
           //------------------------------------------------------------------------------------------
           // Convert relative to absoulte coordinates
           //------------------------------------------------------------------------------------------
           // check for additional circMode = 3 to be activated (LKinLang)
           // Changes CmdType to absolute and converts cirmode 3 to 1
           // --> CmdType = 3 (always absolute as result)
           // --> CircleParameters = calculated arc & updated auxPoint
           IF #pathDataElementPreBuf.cmdParameters.circleParameters.circMode = "LKINCTRL_CIRCMODE_GCODE"
             AND #statSubfunctionStatus = #STATUS_NO_ERROR
           THEN
             #tempRetValWord := "LKinCtrl_ConvCircMode3To1"(coordinates := #pathDataElementPreBuf.cmdCoordinates.absolutePosition,
                                                            lastPos := #statLastPos,
                                                            errorMessage => #statDebugMessage,
                                                            cmdType := #pathDataElementPreBuf.cmdType,
                                                            circleParameters := #pathDataElementPreBuf.cmdParameters.circleParameters);
           END_IF;

           IF #statSubfunctionStatus = #STATUS_NO_ERROR THEN
             // Calculate resulting absoulte position; also convert relative to absolute positions
             #tempRetValWord := "LKinCtrl_CalcResultingPos"(cmdType := #pathDataElementPreBuf.cmdType,
                                                            cartesianPos := #pathDataElementPreBuf.cmdCoordinates.absolutePosition,
                                                            circleParameters := #pathDataElementPreBuf.cmdParameters.circleParameters,
                                                            errorMessage => #statDebugMessage,
                                                            lastAuxPoint := #statAuxPoint, // Absoulte auxPoint
                                                            lastPos := #statLastPos); // Absolute endPoint

             // After this FC call the lastPos equals the endPoint and absolute position
             #statEndPoint := #statAbsolutePosition := #statLastPos;

             // Check if ResultingPos calculation returned an error
             IF #tempRetValWord <> #STATUS_NO_ERROR THEN
               // set error information
               #diagnostics.faultSetNumber := #pathDataElementPreBuf.cmdID;
               #diagnostics.faultPathDataName := #pathDataElementPreBuf.pathDataName;
               #statSubfunctionStatus := #tempRetValWord;
               // set state machine
               #statStateMachine := #ERROR_STATE;
             END_IF;
           END_IF;

         ELSE
           // Command is not a motion command --> WaitTime or FlagOnly
           // ==> Nothing to calculate 
           ;
         END_IF;

         //------------------------------------------------------------------------------------------
         // Command Selection
         //------------------------------------------------------------------------------------------
         // interpretation command to be a linear or circular motion
         IF #statSubfunctionStatus = #STATUS_NO_ERROR THEN
           IF #pathDataElementPreBuf.cmdType = "LKINCTRL_MC_MOVELINEARABS" OR
             #pathDataElementPreBuf.cmdType = "LKINCTRL_MC_MOVELINEARREL" THEN
             #statStateMachine := #EXEC_LIN;
           ELSIF #pathDataElementPreBuf.cmdType = "LKINCTRL_MC_MOVECIRCULARABS" OR
             #pathDataElementPreBuf.cmdType = "LKINCTRL_MC_MOVECIRCULARREL" THEN
             #statStateMachine := #EXEC_CIRC;
           ELSIF #pathDataElementPreBuf.cmdType = "LKINCTRL_MC_MOVEDIRECTABS" OR
             #pathDataElementPreBuf.cmdType = "LKINCTRL_MC_MOVEDIRECTREL" THEN
             #statStateMachine := #EXEC_MOVE_DIRECT;
           ELSIF #pathDataElementPreBuf.cmdType = "LKINCTRL_CMD_WAIT_TIME" THEN
             #statStateMachine := #EXEC_WAIT_TIME;
           ELSIF #pathDataElementPreBuf.cmdType = "LKINCTRL_CMD_FLAG_ONLY" THEN
             #statStateMachine := #EXEC_FLAG_ONLY;
           ELSIF #pathDataElementPreBuf.cmdType = "LKINCTRL_MC_TRACKCONVEYORBELT" THEN
             #statStateMachine := #EXEC_TRACK_CONV;
           END_IF;
         END_IF;
       END_IF;

     END_REGION CMD_CALC 


     // execute MC_MOVELINEARABSOLUTE motion commands  
     REGION EXEC_LIN
       IF #statStateMachine = #EXEC_LIN
         // AND #statDebugState = TRUE
       THEN
         // reset  variable for single step debugging of states
         #statDebugState := FALSE;

         IF #statError = FALSE THEN

           // set execute trigger for linear command
           #statExecLinCmds[#statFBCounterLin] := TRUE;

           // Store motion command data for further calcualtions
           // last position for relative commands
           //#statLastPos := #statAbsolutePosition;

           // command details from PathData and assignment to MC_FBs for activeCmdNo
           #statStoreExecuteBuffer.bufferElement[#statStoreExecuteBuffer.writeBufferElement].pathDataName := #pathDataElementPreBuf.pathDataName;
           #statStoreExecuteBuffer.bufferElement[#statStoreExecuteBuffer.writeBufferElement].pathDataIdentifier := #pathDataElementPreBuf.pathDataIdentifier;
           #statStoreExecuteBuffer.bufferElement[#statStoreExecuteBuffer.writeBufferElement].setNumber := #pathDataElementPreBuf.cmdID;
           #statStoreExecuteBuffer.bufferElement[#statStoreExecuteBuffer.writeBufferElement].MotionFBNo := #statFBCounterLin;
           #statStoreExecuteBuffer.lastBufferElement := #statStoreExecuteBuffer.writeBufferElement;

           // increase writeBufferElement pointer for statStoreBuffer for assignment of activeCmdNo
           IF #statStoreExecuteBuffer.writeBufferElement < #LKINCTRL_EXECUTEBUFFER_LENGTH THEN
             #statStoreExecuteBuffer.writeBufferElement := #statStoreExecuteBuffer.writeBufferElement + 1;
           ELSE
             #statStoreExecuteBuffer.writeBufferElement := 1;
           END_IF;

           REGION CMD_LOGGER
             // // DATA LOGGER handling
             // write command data to data logger
             // single data entries of PathDataElement instead of complete structure ==> to deep nesting level
             #statDebugExecCmdLogger.loggerElement[#statDebugExecCmdLogger.writeCmdLoggerElement].executedCmd.cmdType := #pathDataElementPreBuf.cmdType;
             #statDebugExecCmdLogger.loggerElement[#statDebugExecCmdLogger.writeCmdLoggerElement].executedCmd.pathDataName := #pathDataElementPreBuf.pathDataName;
             #statDebugExecCmdLogger.loggerElement[#statDebugExecCmdLogger.writeCmdLoggerElement].executedCmd.pathDataIdentifier := #pathDataElementPreBuf.pathDataIdentifier;
             #statDebugExecCmdLogger.loggerElement[#statDebugExecCmdLogger.writeCmdLoggerElement].executedCmd.cmdID := #pathDataElementPreBuf.cmdID;
             #statDebugExecCmdLogger.loggerElement[#statDebugExecCmdLogger.writeCmdLoggerElement].executedCmd.cmdName := #pathDataElementPreBuf.cmdName;
             // coordinates logging
             #statDebugExecCmdLogger.loggerElement[#statDebugExecCmdLogger.writeCmdLoggerElement].executedCmd.coordinateX := #pathDataElementPreBuf.cmdCoordinates.absolutePosition[1];
             #statDebugExecCmdLogger.loggerElement[#statDebugExecCmdLogger.writeCmdLoggerElement].executedCmd.coordinateY := #pathDataElementPreBuf.cmdCoordinates.absolutePosition[2];
             #statDebugExecCmdLogger.loggerElement[#statDebugExecCmdLogger.writeCmdLoggerElement].executedCmd.coordinateZ := #pathDataElementPreBuf.cmdCoordinates.absolutePosition[3];
             #statDebugExecCmdLogger.loggerElement[#statDebugExecCmdLogger.writeCmdLoggerElement].executedCmd.coordinateA := #pathDataElementPreBuf.cmdCoordinates.absolutePosition[4];
             #statDebugExecCmdLogger.loggerElement[#statDebugExecCmdLogger.writeCmdLoggerElement].executedCmd.coordSystem := #pathDataElementPreBuf.cmdCoordinates.coordSystem;
             // cmdParameter logging
             #statDebugExecCmdLogger.loggerElement[#statDebugExecCmdLogger.writeCmdLoggerElement].executedCmd.bufferMode := #pathDataElementPreBuf.cmdParameters.bufferMode;
             #statDebugExecCmdLogger.loggerElement[#statDebugExecCmdLogger.writeCmdLoggerElement].executedCmd.transitionParameter := #pathDataElementPreBuf.cmdParameters.transitionParameters[1];
             #statDebugExecCmdLogger.loggerElement[#statDebugExecCmdLogger.writeCmdLoggerElement].executedCmd.dynVelocity := #pathDataElementPreBuf.cmdParameters.pathDynamics.velocity;
             #statDebugExecCmdLogger.loggerElement[#statDebugExecCmdLogger.writeCmdLoggerElement].executedCmd.dynAcceleration := #pathDataElementPreBuf.cmdParameters.pathDynamics.acceleration;
             #statDebugExecCmdLogger.loggerElement[#statDebugExecCmdLogger.writeCmdLoggerElement].executedCmd.dynDeceleration := #pathDataElementPreBuf.cmdParameters.pathDynamics.deceleration;
             #statDebugExecCmdLogger.loggerElement[#statDebugExecCmdLogger.writeCmdLoggerElement].executedCmd.dynJerk := #pathDataElementPreBuf.cmdParameters.pathDynamics.jerk;
             #statDebugExecCmdLogger.loggerElement[#statDebugExecCmdLogger.writeCmdLoggerElement].executedCmd.dynamicAdpation := #pathDataElementPreBuf.cmdParameters.dynamicAdaption;
             // logger element data
             #statDebugExecCmdLogger.loggerElement[#statDebugExecCmdLogger.writeCmdLoggerElement].executeBufferElement := #statStoreExecuteBuffer.lastBufferElement;
             #statDebugExecCmdLogger.loggerElement[#statDebugExecCmdLogger.writeCmdLoggerElement].assignedMotionFB := #statFBCounterLin;
             #tempRetVal := RD_SYS_T(#statDebugExecCmdLogger.loggerElement[#statDebugExecCmdLogger.writeCmdLoggerElement].timeStamp);

             // increment writeCmdLogger pointer
             IF #statDebugExecCmdLogger.writeCmdLoggerElement < #CONST_LENGTH_DATALOGGER THEN
               #statDebugExecCmdLogger.writeCmdLoggerElement := #statDebugExecCmdLogger.writeCmdLoggerElement + 1;
             ELSE
               #statDebugExecCmdLogger.writeCmdLoggerElement := 1;
             END_IF;
           END_REGION CMD_LOGGER

           // set FBCounter variables
           IF #statFBCounterLin < #LKINCTRL_MAX_NUMBER_OF_CMDS_LIN THEN
             #statFBCounterLin := #statFBCounterLin + 1;
           ELSE
             #statFBCounterLin := 1;
           END_IF;

           // set status for outputs
           #statCmdExecuted := TRUE;
           #statStatus := #STATUS_CMD_EXECUTED;

         ELSE
           #statStateMachine := #ERROR_STATE;
         END_IF;
       END_IF;
     END_REGION EXEC_LIN


     // execute MC_MOVECIRCULRABSOLUTE motion commands
     REGION EXEC_CIRC
       IF #statStateMachine = #EXEC_CIRC
         // AND #statDebugState = TRUE
       THEN
         // reset variable for single step debugging of states
         #statDebugState := FALSE;

         IF #statError = FALSE THEN

           // set execute trigger for circular command
           #statExecCircCmds[#statFBCounterCirc] := TRUE;

           // command details from PathData and assignment to MC_FBs for activeCmdNo
           #statStoreExecuteBuffer.bufferElement[#statStoreExecuteBuffer.writeBufferElement].pathDataName := #pathDataElementPreBuf.pathDataName;
           #statStoreExecuteBuffer.bufferElement[#statStoreExecuteBuffer.writeBufferElement].pathDataIdentifier := #pathDataElementPreBuf.pathDataIdentifier;
           #statStoreExecuteBuffer.bufferElement[#statStoreExecuteBuffer.writeBufferElement].setNumber := #pathDataElementPreBuf.cmdID;
           #statStoreExecuteBuffer.bufferElement[#statStoreExecuteBuffer.writeBufferElement].MotionFBNo := #LKINCTRL_EXECUTEBUFFER_LENGTH + #statFBCounterCirc;
           #statStoreExecuteBuffer.lastBufferElement := #statStoreExecuteBuffer.writeBufferElement;

           // increase writeBufferElement pointer for statStoreBuffer for assignment of activeCmdNo
           IF #statStoreExecuteBuffer.writeBufferElement < #LKINCTRL_EXECUTEBUFFER_LENGTH THEN
             #statStoreExecuteBuffer.writeBufferElement := #statStoreExecuteBuffer.writeBufferElement + 1;
           ELSE
             #statStoreExecuteBuffer.writeBufferElement := 1;
           END_IF;

           REGION CMD_LOGGER
             // // DATA LOGGER handling
             // write command data to data logger
             // single data entries of PathDataElement instead of complete structure ==> to deep nesting level
             #statDebugExecCmdLogger.loggerElement[#statDebugExecCmdLogger.writeCmdLoggerElement].executedCmd.cmdType := #pathDataElementPreBuf.cmdType;
             #statDebugExecCmdLogger.loggerElement[#statDebugExecCmdLogger.writeCmdLoggerElement].executedCmd.pathDataName := #pathDataElementPreBuf.pathDataName;
             #statDebugExecCmdLogger.loggerElement[#statDebugExecCmdLogger.writeCmdLoggerElement].executedCmd.pathDataIdentifier := #pathDataElementPreBuf.pathDataIdentifier;
             #statDebugExecCmdLogger.loggerElement[#statDebugExecCmdLogger.writeCmdLoggerElement].executedCmd.cmdID := #pathDataElementPreBuf.cmdID;
             #statDebugExecCmdLogger.loggerElement[#statDebugExecCmdLogger.writeCmdLoggerElement].executedCmd.cmdName := #pathDataElementPreBuf.cmdName;
             // coordinates logging (use auxPoint in X,Y,Z variables)
             #statDebugExecCmdLogger.loggerElement[#statDebugExecCmdLogger.writeCmdLoggerElement].executedCmd.coordinateX := #statEndPoint[1];
             #statDebugExecCmdLogger.loggerElement[#statDebugExecCmdLogger.writeCmdLoggerElement].executedCmd.coordinateY := #statEndPoint[2];
             #statDebugExecCmdLogger.loggerElement[#statDebugExecCmdLogger.writeCmdLoggerElement].executedCmd.coordinateZ := #statEndPoint[3];
             #statDebugExecCmdLogger.loggerElement[#statDebugExecCmdLogger.writeCmdLoggerElement].executedCmd.coordinateA := #statEndPoint[4];
             #statDebugExecCmdLogger.loggerElement[#statDebugExecCmdLogger.writeCmdLoggerElement].executedCmd.coordSystem := #pathDataElementPreBuf.cmdCoordinates.coordSystem;
             // cmdParameter logging
             #statDebugExecCmdLogger.loggerElement[#statDebugExecCmdLogger.writeCmdLoggerElement].executedCmd.bufferMode := #pathDataElementPreBuf.cmdParameters.bufferMode;
             #statDebugExecCmdLogger.loggerElement[#statDebugExecCmdLogger.writeCmdLoggerElement].executedCmd.transitionParameter := #pathDataElementPreBuf.cmdParameters.transitionParameters[1];
             #statDebugExecCmdLogger.loggerElement[#statDebugExecCmdLogger.writeCmdLoggerElement].executedCmd.dynVelocity := #pathDataElementPreBuf.cmdParameters.pathDynamics.velocity;
             #statDebugExecCmdLogger.loggerElement[#statDebugExecCmdLogger.writeCmdLoggerElement].executedCmd.dynAcceleration := #pathDataElementPreBuf.cmdParameters.pathDynamics.acceleration;
             #statDebugExecCmdLogger.loggerElement[#statDebugExecCmdLogger.writeCmdLoggerElement].executedCmd.dynDeceleration := #pathDataElementPreBuf.cmdParameters.pathDynamics.deceleration;
             #statDebugExecCmdLogger.loggerElement[#statDebugExecCmdLogger.writeCmdLoggerElement].executedCmd.dynJerk := #pathDataElementPreBuf.cmdParameters.pathDynamics.jerk;
             #statDebugExecCmdLogger.loggerElement[#statDebugExecCmdLogger.writeCmdLoggerElement].executedCmd.dynamicAdpation := #pathDataElementPreBuf.cmdParameters.dynamicAdaption;
             // circle parameter logging
             #statDebugExecCmdLogger.loggerElement[#statDebugExecCmdLogger.writeCmdLoggerElement].executedCmd.circMode := #pathDataElementPreBuf.cmdParameters.circleParameters.circMode;
             #statDebugExecCmdLogger.loggerElement[#statDebugExecCmdLogger.writeCmdLoggerElement].executedCmd.auxPoint_1 := #pathDataElementPreBuf.cmdParameters.circleParameters.auxPoint[1];
             #statDebugExecCmdLogger.loggerElement[#statDebugExecCmdLogger.writeCmdLoggerElement].executedCmd.auxPoint_2 := #pathDataElementPreBuf.cmdParameters.circleParameters.auxPoint[2];
             #statDebugExecCmdLogger.loggerElement[#statDebugExecCmdLogger.writeCmdLoggerElement].executedCmd.auxPoint_3 := #pathDataElementPreBuf.cmdParameters.circleParameters.auxPoint[3];
             #statDebugExecCmdLogger.loggerElement[#statDebugExecCmdLogger.writeCmdLoggerElement].executedCmd.pathChoice := #pathDataElementPreBuf.cmdParameters.circleParameters.pathChoice;
             #statDebugExecCmdLogger.loggerElement[#statDebugExecCmdLogger.writeCmdLoggerElement].executedCmd.circlePlane := #pathDataElementPreBuf.cmdParameters.circleParameters.circlePlane;
             #statDebugExecCmdLogger.loggerElement[#statDebugExecCmdLogger.writeCmdLoggerElement].executedCmd.radius := #pathDataElementPreBuf.cmdParameters.circleParameters.radius;
             #statDebugExecCmdLogger.loggerElement[#statDebugExecCmdLogger.writeCmdLoggerElement].executedCmd.arc := #pathDataElementPreBuf.cmdParameters.circleParameters.arc;

             // logger element data
             #statDebugExecCmdLogger.loggerElement[#statDebugExecCmdLogger.writeCmdLoggerElement].executeBufferElement := #statStoreExecuteBuffer.lastBufferElement;
             #statDebugExecCmdLogger.loggerElement[#statDebugExecCmdLogger.writeCmdLoggerElement].assignedMotionFB := 10 + #statFBCounterCirc;
             #tempRetVal := RD_SYS_T(#statDebugExecCmdLogger.loggerElement[#statDebugExecCmdLogger.writeCmdLoggerElement].timeStamp);

             // increment writeCmdLogger pointer
             IF #statDebugExecCmdLogger.writeCmdLoggerElement < #CONST_LENGTH_DATALOGGER THEN
               #statDebugExecCmdLogger.writeCmdLoggerElement := #statDebugExecCmdLogger.writeCmdLoggerElement + 1;
             ELSE
               #statDebugExecCmdLogger.writeCmdLoggerElement := 1;
             END_IF;
           END_REGION CMD_LOGGER

           // set FBCounter variables
           IF #statFBCounterCirc < #LKINCTRL_MAX_NUMBER_OF_CMDS_CIRC THEN
             #statFBCounterCirc := #statFBCounterCirc + 1;
           ELSE
             #statFBCounterCirc := 1;
           END_IF;

           // set status for outputs
           #statCmdExecuted := TRUE;
           #statStatus := #STATUS_CMD_EXECUTED;

         ELSE
           #statStateMachine := #ERROR_STATE;
         END_IF;
       END_IF;
     END_REGION EXEC_CIRC


     // execute MC_MOVEDIRECTABSOLUTE motion commands  
     REGION EXEC_MOVE_DIRECT
       IF #statStateMachine = #EXEC_MOVE_DIRECT
         // AND #statDebugState = TRUE
       THEN
         // reset  variable for single step debugging of states
         #statDebugState := FALSE;

         IF #statError = FALSE THEN

           // set execute trigger for move direct command
           #statExecMoveDirectCmds[#statFBCounterMoveDir] := TRUE;

           // Store motion command data for further calcualtions
           // last position for relative commands
           //#statLastPos := #statAbsolutePosition;

           // command details from PathData and assignment to MC_FBs for activeCmdNo
           #statStoreExecuteBuffer.bufferElement[#statStoreExecuteBuffer.writeBufferElement].pathDataName := #pathDataElementPreBuf.pathDataName;
           #statStoreExecuteBuffer.bufferElement[#statStoreExecuteBuffer.writeBufferElement].pathDataIdentifier := #pathDataElementPreBuf.pathDataIdentifier;
           #statStoreExecuteBuffer.bufferElement[#statStoreExecuteBuffer.writeBufferElement].setNumber := #pathDataElementPreBuf.cmdID;
           #statStoreExecuteBuffer.bufferElement[#statStoreExecuteBuffer.writeBufferElement].MotionFBNo := #LKINCTRL_EXECUTEBUFFER_LENGTH + #LKINCTRL_EXECUTEBUFFER_LENGTH + #statFBCounterMoveDir;
           #statStoreExecuteBuffer.lastBufferElement := #statStoreExecuteBuffer.writeBufferElement;

           // increase writeBufferElement pointer for statStoreBuffer for assignment of activeCmdNo
           IF #statStoreExecuteBuffer.writeBufferElement < #LKINCTRL_EXECUTEBUFFER_LENGTH THEN
             #statStoreExecuteBuffer.writeBufferElement := #statStoreExecuteBuffer.writeBufferElement + 1;
           ELSE
             #statStoreExecuteBuffer.writeBufferElement := 1;
           END_IF;

           REGION CMD_LOGGER
             // // DATA LOGGER handling
             // write command data to data logger
             // single data entries of PathDataElement instead of complete structure ==> to deep nesting level
             #statDebugExecCmdLogger.loggerElement[#statDebugExecCmdLogger.writeCmdLoggerElement].executedCmd.cmdType := #pathDataElementPreBuf.cmdType;
             #statDebugExecCmdLogger.loggerElement[#statDebugExecCmdLogger.writeCmdLoggerElement].executedCmd.pathDataName := #pathDataElementPreBuf.pathDataName;
             #statDebugExecCmdLogger.loggerElement[#statDebugExecCmdLogger.writeCmdLoggerElement].executedCmd.pathDataIdentifier := #pathDataElementPreBuf.pathDataIdentifier;
             #statDebugExecCmdLogger.loggerElement[#statDebugExecCmdLogger.writeCmdLoggerElement].executedCmd.cmdID := #pathDataElementPreBuf.cmdID;
             #statDebugExecCmdLogger.loggerElement[#statDebugExecCmdLogger.writeCmdLoggerElement].executedCmd.cmdName := #pathDataElementPreBuf.cmdName;
             // coordinates logging
             #statDebugExecCmdLogger.loggerElement[#statDebugExecCmdLogger.writeCmdLoggerElement].executedCmd.coordinateX := #pathDataElementPreBuf.cmdCoordinates.absolutePosition[1];
             #statDebugExecCmdLogger.loggerElement[#statDebugExecCmdLogger.writeCmdLoggerElement].executedCmd.coordinateY := #pathDataElementPreBuf.cmdCoordinates.absolutePosition[2];
             #statDebugExecCmdLogger.loggerElement[#statDebugExecCmdLogger.writeCmdLoggerElement].executedCmd.coordinateZ := #pathDataElementPreBuf.cmdCoordinates.absolutePosition[3];
             #statDebugExecCmdLogger.loggerElement[#statDebugExecCmdLogger.writeCmdLoggerElement].executedCmd.coordinateA := #pathDataElementPreBuf.cmdCoordinates.absolutePosition[4];
             #statDebugExecCmdLogger.loggerElement[#statDebugExecCmdLogger.writeCmdLoggerElement].executedCmd.coordSystem := #pathDataElementPreBuf.cmdCoordinates.coordSystem;
             // cmdParameter logging
             #statDebugExecCmdLogger.loggerElement[#statDebugExecCmdLogger.writeCmdLoggerElement].executedCmd.bufferMode := #pathDataElementPreBuf.cmdParameters.bufferMode;
             #statDebugExecCmdLogger.loggerElement[#statDebugExecCmdLogger.writeCmdLoggerElement].executedCmd.transitionParameter := #pathDataElementPreBuf.cmdParameters.transitionParameters[1];
             #statDebugExecCmdLogger.loggerElement[#statDebugExecCmdLogger.writeCmdLoggerElement].executedCmd.dynVelocity := #pathDataElementPreBuf.cmdParameters.pathDynamics.velocity;
             #statDebugExecCmdLogger.loggerElement[#statDebugExecCmdLogger.writeCmdLoggerElement].executedCmd.dynAcceleration := #pathDataElementPreBuf.cmdParameters.pathDynamics.acceleration;
             #statDebugExecCmdLogger.loggerElement[#statDebugExecCmdLogger.writeCmdLoggerElement].executedCmd.dynDeceleration := #pathDataElementPreBuf.cmdParameters.pathDynamics.deceleration;
             #statDebugExecCmdLogger.loggerElement[#statDebugExecCmdLogger.writeCmdLoggerElement].executedCmd.dynJerk := #pathDataElementPreBuf.cmdParameters.pathDynamics.jerk;
             #statDebugExecCmdLogger.loggerElement[#statDebugExecCmdLogger.writeCmdLoggerElement].executedCmd.dynamicAdpation := #pathDataElementPreBuf.cmdParameters.dynamicAdaption;

             #statDebugExecCmdLogger.loggerElement[#statDebugExecCmdLogger.writeCmdLoggerElement].executedCmd.linkConstellation := #pathDataElementPreBuf.cmdParameters.moveDirectParameters.linkConstellation;
             #statDebugExecCmdLogger.loggerElement[#statDebugExecCmdLogger.writeCmdLoggerElement].executedCmd.positionMode := #pathDataElementPreBuf.cmdParameters.moveDirectParameters.positionMode;

             // logger element data
             #statDebugExecCmdLogger.loggerElement[#statDebugExecCmdLogger.writeCmdLoggerElement].executeBufferElement := #statStoreExecuteBuffer.lastBufferElement;
             #statDebugExecCmdLogger.loggerElement[#statDebugExecCmdLogger.writeCmdLoggerElement].assignedMotionFB := #statFBCounterMoveDir;
             #tempRetVal := RD_SYS_T(#statDebugExecCmdLogger.loggerElement[#statDebugExecCmdLogger.writeCmdLoggerElement].timeStamp);

             // increment writeCmdLogger pointer
             IF #statDebugExecCmdLogger.writeCmdLoggerElement < #CONST_LENGTH_DATALOGGER THEN
               #statDebugExecCmdLogger.writeCmdLoggerElement := #statDebugExecCmdLogger.writeCmdLoggerElement + 1;
             ELSE
               #statDebugExecCmdLogger.writeCmdLoggerElement := 1;
             END_IF;
           END_REGION CMD_LOGGER

           // set FBCounter variables
           IF #statFBCounterMoveDir < #LKINCTRL_MAX_NUMBER_OF_CMDS_MOVEDIRECT THEN
             #statFBCounterMoveDir := #statFBCounterMoveDir + 1;
           ELSE
             #statFBCounterMoveDir := 1;
           END_IF;

           // set status for outputs
           #statCmdExecuted := TRUE;
           #statStatus := #STATUS_CMD_EXECUTED;

         ELSE
           #statStateMachine := #ERROR_STATE;
         END_IF;
       END_IF;
     END_REGION EXEC_MOVE_DIRECT


     // execute MC_TRACKCONVEYORBELT motion commands  
     REGION EXEC_TRACK_CONVEYOR
       IF #statStateMachine = #EXEC_TRACK_CONV
         // AND #statDebugState = TRUE
       THEN
         // reset  variable for single step debugging of states
         #statDebugState := FALSE;

         IF #statError = FALSE THEN

           // set execute trigger for move direct command
           #statExecTrackConv[#statFBCounterTrackConv] := TRUE;

           // Copy conveyor configuration to instance
           #statConveyorBeltAxis[#statFBCounterTrackConv] := #conveyorConfiguration[#pathDataElementPreBuf.cmdParameters.conveyorParameters.conveyorParaNo].conveyorBeltAxis;
           #instMC_TrackConveyor[#statFBCounterTrackConv].ConveyorBeltOrigin := #conveyorConfiguration[#pathDataElementPreBuf.cmdParameters.conveyorParameters.conveyorParaNo].conveyorBeltOrigin;
           #instMC_TrackConveyor[#statFBCounterTrackConv].InitialObjectPosition := #conveyorConfiguration[#pathDataElementPreBuf.cmdParameters.conveyorParameters.conveyorParaNo].initialObjectPosition;
           #instMC_TrackConveyor[#statFBCounterTrackConv].CoordSystem := #pathDataElementPreBuf.cmdCoordinates.coordSystem;

           // Set OCS in tracking
           #statOCSInTracking[#instMC_TrackConveyor[#statFBCounterTrackConv].CoordSystem] := TRUE;

           // command details from PathData and assignment to MC_FBs for activeCmdNo
           #statStoreExecuteBuffer.bufferElement[#statStoreExecuteBuffer.writeBufferElement].pathDataName := #pathDataElementPreBuf.pathDataName;
           #statStoreExecuteBuffer.bufferElement[#statStoreExecuteBuffer.writeBufferElement].pathDataIdentifier := #pathDataElementPreBuf.pathDataIdentifier;
           #statStoreExecuteBuffer.bufferElement[#statStoreExecuteBuffer.writeBufferElement].setNumber := #pathDataElementPreBuf.cmdID;
           #statStoreExecuteBuffer.bufferElement[#statStoreExecuteBuffer.writeBufferElement].MotionFBNo := "LKINCTRL_CMD_WAIT_TIME" + #statFBCounterTrackConv;
           #statStoreExecuteBuffer.lastBufferElement := #statStoreExecuteBuffer.writeBufferElement;

           // increase writeBufferElement pointer for statStoreBuffer for assignment of activeCmdNo
           IF #statStoreExecuteBuffer.writeBufferElement < #LKINCTRL_EXECUTEBUFFER_LENGTH THEN
             #statStoreExecuteBuffer.writeBufferElement := #statStoreExecuteBuffer.writeBufferElement + 1;
           ELSE
             #statStoreExecuteBuffer.writeBufferElement := 1;
           END_IF;

           REGION CMD_LOGGER
             // // DATA LOGGER handling
             // write command data to data logger
             // single data entries of PathDataElement instead of complete structure ==> to deep nesting level
             #statDebugExecCmdLogger.loggerElement[#statDebugExecCmdLogger.writeCmdLoggerElement].executedCmd.cmdType := #pathDataElementPreBuf.cmdType;
             #statDebugExecCmdLogger.loggerElement[#statDebugExecCmdLogger.writeCmdLoggerElement].executedCmd.pathDataName := #pathDataElementPreBuf.pathDataName;
             #statDebugExecCmdLogger.loggerElement[#statDebugExecCmdLogger.writeCmdLoggerElement].executedCmd.pathDataIdentifier := #pathDataElementPreBuf.pathDataIdentifier;
             #statDebugExecCmdLogger.loggerElement[#statDebugExecCmdLogger.writeCmdLoggerElement].executedCmd.cmdID := #pathDataElementPreBuf.cmdID;
             #statDebugExecCmdLogger.loggerElement[#statDebugExecCmdLogger.writeCmdLoggerElement].executedCmd.cmdName := #pathDataElementPreBuf.cmdName;
             // coordinates logging
             #statDebugExecCmdLogger.loggerElement[#statDebugExecCmdLogger.writeCmdLoggerElement].executedCmd.coordinateX := #pathDataElementPreBuf.cmdCoordinates.absolutePosition[1];
             #statDebugExecCmdLogger.loggerElement[#statDebugExecCmdLogger.writeCmdLoggerElement].executedCmd.coordinateY := #pathDataElementPreBuf.cmdCoordinates.absolutePosition[2];
             #statDebugExecCmdLogger.loggerElement[#statDebugExecCmdLogger.writeCmdLoggerElement].executedCmd.coordinateZ := #pathDataElementPreBuf.cmdCoordinates.absolutePosition[3];
             #statDebugExecCmdLogger.loggerElement[#statDebugExecCmdLogger.writeCmdLoggerElement].executedCmd.coordinateA := #pathDataElementPreBuf.cmdCoordinates.absolutePosition[4];
             #statDebugExecCmdLogger.loggerElement[#statDebugExecCmdLogger.writeCmdLoggerElement].executedCmd.coordSystem := #pathDataElementPreBuf.cmdCoordinates.coordSystem;
             // cmdParameter logging
             #statDebugExecCmdLogger.loggerElement[#statDebugExecCmdLogger.writeCmdLoggerElement].executedCmd.bufferMode := #pathDataElementPreBuf.cmdParameters.bufferMode;
             #statDebugExecCmdLogger.loggerElement[#statDebugExecCmdLogger.writeCmdLoggerElement].executedCmd.transitionParameter := #pathDataElementPreBuf.cmdParameters.transitionParameters[1];
             #statDebugExecCmdLogger.loggerElement[#statDebugExecCmdLogger.writeCmdLoggerElement].executedCmd.dynVelocity := #pathDataElementPreBuf.cmdParameters.pathDynamics.velocity;
             #statDebugExecCmdLogger.loggerElement[#statDebugExecCmdLogger.writeCmdLoggerElement].executedCmd.dynAcceleration := #pathDataElementPreBuf.cmdParameters.pathDynamics.acceleration;
             #statDebugExecCmdLogger.loggerElement[#statDebugExecCmdLogger.writeCmdLoggerElement].executedCmd.dynDeceleration := #pathDataElementPreBuf.cmdParameters.pathDynamics.deceleration;
             #statDebugExecCmdLogger.loggerElement[#statDebugExecCmdLogger.writeCmdLoggerElement].executedCmd.dynJerk := #pathDataElementPreBuf.cmdParameters.pathDynamics.jerk;
             #statDebugExecCmdLogger.loggerElement[#statDebugExecCmdLogger.writeCmdLoggerElement].executedCmd.dynamicAdpation := #pathDataElementPreBuf.cmdParameters.dynamicAdaption;

             #statDebugExecCmdLogger.loggerElement[#statDebugExecCmdLogger.writeCmdLoggerElement].executedCmd.linkConstellation := #pathDataElementPreBuf.cmdParameters.moveDirectParameters.linkConstellation;
             #statDebugExecCmdLogger.loggerElement[#statDebugExecCmdLogger.writeCmdLoggerElement].executedCmd.positionMode := #pathDataElementPreBuf.cmdParameters.moveDirectParameters.positionMode;

             // logger element data
             #statDebugExecCmdLogger.loggerElement[#statDebugExecCmdLogger.writeCmdLoggerElement].executeBufferElement := #statStoreExecuteBuffer.lastBufferElement;
             #statDebugExecCmdLogger.loggerElement[#statDebugExecCmdLogger.writeCmdLoggerElement].assignedMotionFB := #statFBCounterTrackConv;
             #tempRetVal := RD_SYS_T(#statDebugExecCmdLogger.loggerElement[#statDebugExecCmdLogger.writeCmdLoggerElement].timeStamp);

             // increment writeCmdLogger pointer
             IF #statDebugExecCmdLogger.writeCmdLoggerElement < #CONST_LENGTH_DATALOGGER THEN
               #statDebugExecCmdLogger.writeCmdLoggerElement := #statDebugExecCmdLogger.writeCmdLoggerElement + 1;
             ELSE
               #statDebugExecCmdLogger.writeCmdLoggerElement := 1;
             END_IF;
           END_REGION CMD_LOGGER

           // set FBCounter variables
           IF #statFBCounterTrackConv < #LKINCTRL_MAX_NUMBER_OF_CMDS_TRACKCONV THEN
             #statFBCounterTrackConv := #statFBCounterTrackConv + 1;
           ELSE
             #statFBCounterTrackConv := 1;
           END_IF;

           // set status for outputs
           #statCmdExecuted := TRUE;
           #statStatus := #STATUS_CMD_EXECUTED;

         ELSE
           #statStateMachine := #ERROR_STATE;
         END_IF;
       END_IF;
     END_REGION EXEC_TRACK_CONVEYOR



     // execute WAIT TIME 
     REGION EXEC_WAIT_TIME
       IF #statStateMachine = #EXEC_WAIT_TIME
         // AND #statDebugState = TRUE
       THEN
         // reset  variable for single step debugging of states
         #statDebugState := FALSE;

         // check for error to be pending
         IF #statError = FALSE THEN

           // Added check for active mc command; FR: 27.05.2019
           // check for active MC linear instance
           FOR #tempCtr := 1 TO #LKINCTRL_MAX_NUMBER_OF_CMDS_LIN DO
             IF #instMC_MoveLinAbs[#tempCtr].Busy THEN
               // set temp to interlock reset
               #tempMCActive := TRUE;
               EXIT;
             ELSE
               #tempMCActive := FALSE;
             END_IF;
           END_FOR;

           // check for no circular instance to be busy in case of no linear cmd busy
           IF #tempMCActive = FALSE THEN
             FOR #tempCtr := 1 TO #LKINCTRL_MAX_NUMBER_OF_CMDS_CIRC DO
               IF #instMC_MoveCircAbs[#tempCtr].Busy THEN
                 // set temp to interlock reset
                 #tempMCActive := TRUE;
                 EXIT;
               ELSE
                 #tempMCActive := FALSE;
               END_IF;
             END_FOR;
           END_IF;

           // check for no PTP instance to be busy in case of no linear cmd busy
           IF #tempMCActive = FALSE THEN
             FOR #tempCtr := 1 TO #LKINCTRL_MAX_NUMBER_OF_CMDS_MOVEDIRECT DO
               IF #instMC_MoveDirectAbs[#tempCtr].Busy THEN
                 // set temp to interlock reset
                 #tempMCActive := TRUE;
                 EXIT;
               ELSE
                 #tempMCActive := FALSE;
               END_IF;
             END_FOR;
           END_IF;

           // check for previously executed commands to be finished
           IF #to_Kinematics.StatusMotionQueue.NumberOfCommands = 0
             AND #statActive = FALSE
             AND #tempMCActive = FALSE
           THEN
             // read wait time - duration [ms]
             #statWaitTime := INT_TO_TIME(LREAL_TO_INT(#pathDataElementPreBuf.cmdParameters.pathDynamics.velocity));

             // set execute trigger to run timer
             #statExecWaitTime := TRUE;

             // command details from PathData and assignment to MC_FBs for activeCmdNo
             #statStoreExecuteBuffer.bufferElement[#statStoreExecuteBuffer.writeBufferElement].pathDataName := #pathDataElementPreBuf.pathDataName;
             #statStoreExecuteBuffer.bufferElement[#statStoreExecuteBuffer.writeBufferElement].pathDataIdentifier := #pathDataElementPreBuf.pathDataIdentifier;
             #statStoreExecuteBuffer.bufferElement[#statStoreExecuteBuffer.writeBufferElement].setNumber := #pathDataElementPreBuf.cmdID;
             #statStoreExecuteBuffer.bufferElement[#statStoreExecuteBuffer.writeBufferElement].MotionFBNo := "LKINCTRL_CMD_WAIT_TIME";
             #statStoreExecuteBuffer.lastBufferElement := #statStoreExecuteBuffer.writeBufferElement;

             // increase writeBufferElement pointer for statStoreBuffer for assignment of activeCmdNo
             IF #statStoreExecuteBuffer.writeBufferElement < #LKINCTRL_EXECUTEBUFFER_LENGTH THEN
               #statStoreExecuteBuffer.writeBufferElement := #statStoreExecuteBuffer.writeBufferElement + 1;
             ELSE
               #statStoreExecuteBuffer.writeBufferElement := 1;
             END_IF;

             REGION CMD_LOGGER
               // // DATA LOGGER handling
               // write command data to data logger
               // single data entries of PathDataElement instead of complete structure ==> to deep nesting level
               #statDebugExecCmdLogger.loggerElement[#statDebugExecCmdLogger.writeCmdLoggerElement].executedCmd.cmdType := #pathDataElementPreBuf.cmdType;
               #statDebugExecCmdLogger.loggerElement[#statDebugExecCmdLogger.writeCmdLoggerElement].executedCmd.pathDataName := #pathDataElementPreBuf.pathDataName;
               #statDebugExecCmdLogger.loggerElement[#statDebugExecCmdLogger.writeCmdLoggerElement].executedCmd.pathDataIdentifier := #pathDataElementPreBuf.pathDataIdentifier;
               #statDebugExecCmdLogger.loggerElement[#statDebugExecCmdLogger.writeCmdLoggerElement].executedCmd.cmdID := #pathDataElementPreBuf.cmdID;
               #statDebugExecCmdLogger.loggerElement[#statDebugExecCmdLogger.writeCmdLoggerElement].executedCmd.cmdName := #pathDataElementPreBuf.cmdName;
               // parameter logging
               #statDebugExecCmdLogger.loggerElement[#statDebugExecCmdLogger.writeCmdLoggerElement].executedCmd.dynVelocity := #pathDataElementPreBuf.cmdParameters.pathDynamics.velocity;
               // logger element data
               #statDebugExecCmdLogger.loggerElement[#statDebugExecCmdLogger.writeCmdLoggerElement].executeBufferElement := #statStoreExecuteBuffer.lastBufferElement;
               #statDebugExecCmdLogger.loggerElement[#statDebugExecCmdLogger.writeCmdLoggerElement].assignedMotionFB := "LKINCTRL_CMD_WAIT_TIME";
               #tempRetVal := RD_SYS_T(#statDebugExecCmdLogger.loggerElement[#statDebugExecCmdLogger.writeCmdLoggerElement].timeStamp);

               // increment writeCmdLogger pointer
               IF #statDebugExecCmdLogger.writeCmdLoggerElement < #CONST_LENGTH_DATALOGGER THEN
                 #statDebugExecCmdLogger.writeCmdLoggerElement := #statDebugExecCmdLogger.writeCmdLoggerElement + 1;
               ELSE
                 #statDebugExecCmdLogger.writeCmdLoggerElement := 1;
               END_IF;
             END_REGION CMD_LOGGER

             // set cmdExecuted
             #statCmdExecuted := TRUE;
             // set state to signalize WAIT_TIME running
             #statStatus := #STATUS_WAIT_TIME_ACTIVE;
             // go to state to wait for WAIT_TIME to finish
             #statStateMachine := #WAITING_TIME;
           END_IF;

         ELSE
           #statStateMachine := #ERROR_STATE;
         END_IF;
       END_IF;
     END_REGION EXEC_WAIT_TIME


     // execute FLAG_ONLY commands  
     REGION EXEC_FLAG_ONLY
       IF #statStateMachine = #EXEC_FLAG_ONLY
         // AND #statDebugState = TRUE
       THEN
         // reset  variable for single step debugging of states
         #statDebugState := FALSE;

         IF #statError = FALSE THEN

           // checked for PathData to start with flagOnly command in the triggering section (must not be 1st command)
           // set flagOnlyCmd bit manually, as no previous MC command will be 'done' before

           IF #statStartCmdIsFlagOnly THEN
             // set execute trigger here only when PathData starts with flagOnly command
             #statExecuteFlagOnlyCmd := TRUE;
             // reset bit to recognize FlagOnly command
             #statStartCmdIsFlagOnly := FALSE;
           END_IF;

           // command details from PathData and assignment to MC_FBs for activeCmdNo
           #statStoreExecuteBuffer.bufferElement[#statStoreExecuteBuffer.writeBufferElement].pathDataName := #pathDataElementPreBuf.pathDataName;
           #statStoreExecuteBuffer.bufferElement[#statStoreExecuteBuffer.writeBufferElement].pathDataIdentifier := #pathDataElementPreBuf.pathDataIdentifier;
           #statStoreExecuteBuffer.bufferElement[#statStoreExecuteBuffer.writeBufferElement].setNumber := #pathDataElementPreBuf.cmdID;
           #statStoreExecuteBuffer.bufferElement[#statStoreExecuteBuffer.writeBufferElement].MotionFBNo := "LKINCTRL_CMD_FLAG_ONLY";
           #statStoreExecuteBuffer.lastBufferElement := #statStoreExecuteBuffer.writeBufferElement;

           // increase writeBufferElement pointer for statStoreBuffer for assignment of activeCmdNo
           IF #statStoreExecuteBuffer.writeBufferElement < #LKINCTRL_EXECUTEBUFFER_LENGTH THEN
             #statStoreExecuteBuffer.writeBufferElement := #statStoreExecuteBuffer.writeBufferElement + 1;
           ELSE
             #statStoreExecuteBuffer.writeBufferElement := 1;
           END_IF;

           REGION CMD_LOGGER
             // // DATA LOGGER handling
             // write command data to data logger
             // single data entries of PathDataElement instead of complete structure ==> to deep nesting level
             #statDebugExecCmdLogger.loggerElement[#statDebugExecCmdLogger.writeCmdLoggerElement].executedCmd.cmdType := #pathDataElementPreBuf.cmdType;
             #statDebugExecCmdLogger.loggerElement[#statDebugExecCmdLogger.writeCmdLoggerElement].executedCmd.pathDataName := #pathDataElementPreBuf.pathDataName;
             #statDebugExecCmdLogger.loggerElement[#statDebugExecCmdLogger.writeCmdLoggerElement].executedCmd.pathDataIdentifier := #pathDataElementPreBuf.pathDataIdentifier;
             #statDebugExecCmdLogger.loggerElement[#statDebugExecCmdLogger.writeCmdLoggerElement].executedCmd.cmdID := #pathDataElementPreBuf.cmdID;
             #statDebugExecCmdLogger.loggerElement[#statDebugExecCmdLogger.writeCmdLoggerElement].executedCmd.cmdName := #pathDataElementPreBuf.cmdName;

             // logger element data
             #statDebugExecCmdLogger.loggerElement[#statDebugExecCmdLogger.writeCmdLoggerElement].executeBufferElement := #statStoreExecuteBuffer.lastBufferElement;
             #statDebugExecCmdLogger.loggerElement[#statDebugExecCmdLogger.writeCmdLoggerElement].assignedMotionFB := "LKINCTRL_CMD_FLAG_ONLY";
             #tempRetVal := RD_SYS_T(#statDebugExecCmdLogger.loggerElement[#statDebugExecCmdLogger.writeCmdLoggerElement].timeStamp);

             // increment writeCmdLogger pointer
             IF #statDebugExecCmdLogger.writeCmdLoggerElement < #CONST_LENGTH_DATALOGGER THEN
               #statDebugExecCmdLogger.writeCmdLoggerElement := #statDebugExecCmdLogger.writeCmdLoggerElement + 1;
             ELSE
               #statDebugExecCmdLogger.writeCmdLoggerElement := 1;
             END_IF;
           END_REGION CMD_LOGGER

           // set status for outputs
           #statCmdExecuted := TRUE;
           #statStatus := #STATUS_CMD_EXECUTED;

         ELSE
           #statStateMachine := #ERROR_STATE;
         END_IF;
       END_IF;
     END_REGION EXEC_FLAG_ONLY


     // wait for WAIT_TIME to finish
     REGION WAITING_TIME
       IF #statStateMachine = #WAITING_TIME
         // AND #statDebugState = TRUE
       THEN
         // reset  variable for single step debugging of states
         #statDebugState := FALSE;

         // Set waitTimeActive output
         #statWaitTimeActive := TRUE;

         IF #instIEC_Timer_waitTime.Q THEN
           // reset timer by calling with false
           #statExecWaitTime := FALSE;

           // set status for outputs only after time is done
           #statCmdExecuted := TRUE;

           // Reset output
           #statWaitTimeActive := FALSE;

           #statStatus := #STATUS_WAIT_TIME_FINISHED;
         END_IF;

       END_IF;
     END_REGION WAITING_TIME


     // state reached when GroupInterrupt is interrupted ==> do nothing when interrupted
     REGION CONTINUEING 
       IF #statStateMachine = #CONTINUEING
         // AND #statDebugState = TRUE
       THEN
         // reset  variable for single step debugging of states
         #statDebugState := FALSE;

         // check for MC_GroupContinue to be performed successfully  (TO Kinematics not interrupted anymore)
         IF #to_Kinematics.StatusWord.%X17 = FALSE THEN
           #statStateMachine := #CONTINUED;
         ELSE // Added FR 2019/04/12
           // execute MC_GroupContinue only when kinematics is interrupted
           #statExecGroupContinue := TRUE;
         END_IF;

       END_IF;
     END_REGION CONTINUEING


     // state reached when GroupContinue is done ==> do nothing when path motion continues
     REGION CONTINUED
       IF #statStateMachine = #CONTINUED
         // AND #statDebugState = TRUE
       THEN
         // reset  variable for single step debugging of states
         #statDebugState := FALSE;

         IF #instMC_GROUPCONTINUE.Done OR #to_Kinematics.StatusWord.%X17 = FALSE THEN // Also check X17 to be false in case of no GroupContinue // FR 2019/04/12
           // action after continue tbd
           #statStatus := #STATUS_PATHMOTION_RUNNING;
         END_IF;
         // reset execute of MC_GroupContinue when GroupContinue has been triggered
         #statExecGroupContinue := FALSE;

         // FR 11.03.2020: Continue during waitTime --> Start timer again and set state machine to correct state
         IF #statWaitTimeActive THEN
           #statExecWaitTime := TRUE;
           #statStateMachine := #WAITING_TIME;
         END_IF;


       END_IF;
     END_REGION MOTION_CONTINUED


     // state reached to execute MC_GroupInterrupt ==> wait for interrupt to be done
     REGION INTERRUPTING
       IF #statStateMachine = #INTERRUPTING
         // AND #statDebugState = TRUE
       THEN
         // reset  variable for single step debugging of states
         #statDebugState := FALSE;

         // FR 11.03.2020: Interrupt during waitTime --> Save remaining time and stop timer
         IF #statWaitTimeActive THEN
           #statWaitTime := #instIEC_Timer_waitTime.PT - #instIEC_Timer_waitTime.ET;
           #statExecWaitTime := FALSE;
         END_IF;

         // FR 25.06.2020:
         // Kinematics now always shows X17 regardless of active command 
         // --> Changed condition to only check X17
         // --> old code is below
         // check for MC_GroupInterrupt to be completed successfully
         IF #instMC_GROUPCONTINUE.Busy THEN // continue is running and interupt is triggered 
           #statExecGroupContinue := FALSE;
           #statExecGroupInterrupt := TRUE;
         ELSIF #to_Kinematics.StatusWord.%X17 THEN
           #statStateMachine := #INTERRUPTED;
           #statStatus := #STATUS_PATHMOTION_INTERRUPTED;
           #statExecGroupInterrupt := FALSE;
         ELSE
           // execute MC_GroupInterrupt if not already executed or done
           #statExecGroupInterrupt := TRUE;
         END_IF;

         // Old code
         (* IF #instMC_GROUPINTERRUPT.Busy = FALSE THEN
                   // check for MC_GroupInterrupt to be completed successfully
                   IF #to_Kinematics.StatusWord.%X17
                       // Added FR 2019/04/12: If no motionCmd active go to interrupted
                       OR (#to_Kinematics.StatusWord.%X6
                       AND #to_Kinematics.StatusWord.%X12
                       AND #to_Kinematics.StatusPath.Velocity = 0.0
                       AND #to_Kinematics.StatusMotionQueue.NumberOfCommands = 0)
                   THEN
                       #statStateMachine := #INTERRUPTED;
                       #statStatus := #STATUS_PATHMOTION_INTERRUPTED;
                   ELSE
                       // execute MC_GroupInterrupt if not already executed or done
                       #statExecGroupInterrupt := TRUE;
                   END_IF;
               ELSE
                   // reset execute of MC_Groupinterrupt when GroupInterrupt has been triggered
                   #statExecGroupInterrupt := FALSE;
               END_IF; *)

       END_IF;
     END_REGION INTERRUPTING


     // state reached when GroupInterrupt is done ==> do nothing when interrupted
     REGION INTERRUPTED
       IF #statStateMachine = #INTERRUPTED
         // AND #statDebugState = TRUE
       THEN
         // reset  variable for single step debugging of states
         #statDebugState := FALSE;

         // do nothing
         ;
       END_IF;
     END_REGION INTERRUPTED


     // state reached to execute MC_GroupStop ==> wait for stop to be done
     REGION STOPPING
       IF #statStateMachine = #STOPPING
         // AND #statDebugState = TRUE
       THEN
         // reset  variable for single step debugging of states
         #statDebugState := FALSE;

         // reset all execute triggers for motion commands in case of STOP
         FOR #tempCtr := 1 TO #LKINCTRL_MAX_NUMBER_OF_CMDS_LIN DO
           #statExecLinCmds[#tempCtr] := FALSE;
           #statExecCircCmds[#tempCtr] := FALSE;
           #statExecMoveDirectCmds[#tempCtr] := FALSE;
         END_FOR;

         FOR #tempCtr := 1 TO #LKINCTRL_MAX_NUMBER_OF_CMDS_TRACKCONV DO
           #statExecTrackConv[#tempCtr] := FALSE;
         END_FOR;

         // Deactivate waitTime
         #statExecWaitTime := FALSE;
         #statWaitTime := t#0s;

         // set status accordingly
         #statStatus := #STATUS_PATHMOTION_STOPPING;

